           // ******************************************************************************************************
       2: // Start Movement via Processchannel
           // Mode 04 hex = Profile Velocity (RefA32 = target velocity / RefB32 = reserved)
           #ILx2T_Ref.q_dw_refB_32 := 0;
           #ILx2T_Ref.q_dw_refA_16 := INT_TO_WORD(#i_inTargetVelocity);
           #inTargetVelocityHelper := #i_inTargetVelocity;
           #ILx2T_Ref.q_wo_dmControl := #ILx2T_Ref.q_wo_dmControl AND 16#FF80;
           #ILx2T_Ref.q_wo_dmControl := #ILx2T_Ref.q_wo_dmControl OR 16#0004;
           #inState := #inState + 1;
           // ******************************************************************************************************
       3: // Mode Toggle
           #xModeToggleHelper := NOT #ILx2T_Ref.st_ModeStatus.ModeToggle;   // save toggle bit 
           IF NOT #xModeToggleHelper THEN
               #ILx2T_Ref.q_wo_dmControl := #ILx2T_Ref.q_wo_dmControl AND 16#FF7F;
           ELSE
               #ILx2T_Ref.q_wo_dmControl := #ILx2T_Ref.q_wo_dmControl OR 16#0080;
           END_IF;
           #inState := #inState + 1;
           // ******************************************************************************************************
       4: // Check for mode response OK
           // Check for mode toggle and number of operating mode OK
           IF NOT (#xModeToggleHelper XOR #ILx2T_Ref.st_ModeStatus.ModeToggle) AND (#ILx2T_Ref.by_OP_ModeAct = 16#0004) THEN                            // Check operating mode number
               #TON_Timeout(IN := FALSE,
                            PT := t#1s);
               #inState := #inState + 1;
           ELSE
               // TIMEOUT ERROR
               #TON_Timeout(IN := TRUE,
                            PT := t#1s);
               IF #TON_Timeout.Q THEN
                   #TON_Timeout(IN := FALSE,
                                PT := t#1s);
                   #q_xError := TRUE;
                   #inErrorState := #inState;
                   #inState := 100;
               END_IF;
           END_IF;
           // ******************************************************************************************************
       5: // Check operating mode
           // Check for target reached (Drive status x_Add)
           IF (#ILx2T_Ref.i_woDriveStatus AND 16#2000) = 16#2000 THEN  // x_Add = Target vel reached     
               #q_xTargetVelocityReached := TRUE;
           ELSE
               #q_xTargetVelocityReached := FALSE;
           END_IF;
           // x_Error
           IF (#ILx2T_Ref.i_woDriveStatus AND 16#8000) = 16#8000 THEN  // error     
               #inErrorState := #inState;
               #inState := 100;
           // Monitoring of actual operating mode
           ELSIF (#ILx2T_Ref.by_OP_ModeAct <> 16#0004) THEN
               #q_xCommandAborted := TRUE;
               #q_xBusy := FALSE;
               #q_xTargetVelocityReached := FALSE;
               #inState := 110;
           // Check for new target velocity value !
           ELSIF #inTargetVelocityHelper <> #i_inTargetVelocity THEN
               #inState := 2;
           // Check for ABORT command
           ELSIF #i_xAbort THEN
               #ILx2T_Ref.x_QuickStopInt := TRUE;
               #inState := #inState + 1;
           END_IF;
       6:
           #TON_Timeout(IN := TRUE,
                        PT := t#10s);
           IF #TON_Timeout.Q THEN
               #TON_Timeout(IN := FALSE,
                            PT := t#1s);
               #ILx2T_Ref.x_QuickStopInt := FALSE;
               #ILx2T_Ref.x_FaultResetInt := FALSE;
               #q_xError := TRUE;
               #inErrorState := #inState;
               #inState := 100;
           ELSIF #ILx2T_Ref.stDriveStatus.x_End AND (#ILx2T_Ref.i_woDriveStatus AND 16#F) >= 7 THEN  // Check for STANDSTILL
               #ILx2T_Ref.x_QuickStopInt := FALSE;
               #ILx2T_Ref.x_FaultResetInt := TRUE;
           ELSIF #ILx2T_Ref.stDriveStatus.x_End AND (#ILx2T_Ref.i_woDriveStatus AND 16#F) < 7 THEN  // Check for STANDSTILL
               #TON_Timeout(IN := FALSE,
                            PT := t#1s);
               #ILx2T_Ref.x_QuickStopInt := FALSE;
               #ILx2T_Ref.x_FaultResetInt := FALSE;
               #q_xCommandAborted := TRUE;
               #q_xBusy := FALSE;
               #q_xTargetVelocityReached := FALSE;
               #inState := 110;
           END_IF;

           // ******************************************************************************************************
       100:  // Error state
           #q_xBusy := FALSE;
           #q_xError := TRUE;
           #inState := 110;
           // ******************************************************************************************************
       110:  // finished
           IF NOT #i_xExecute AND NOT #i_xAbort THEN
               #q_xTargetVelocityReached := FALSE;
               #q_xError := FALSE;
               #q_xBusy := FALSE;
               #q_xCommandAborted := FALSE;
               #inState := 0;
           END_IF;
           // ******************************************************************************************************
   END_CASE;
END_FUNCTION_BLOCK

FUNCTION_BLOCK "ILx2_ModbusTCP_Data_1500"   // FB10, SCL
{ S7_Optimized_Access := 'FALSE' }
VERSION : 1.5
   VAR_INPUT
      CONNECT_ID_1 : Conn_Ouc := 1;   // unique connection ID DPL Read
      CONNECT_ID_2 : Conn_Ouc := 2;   // unique connection ID DPL Write
      CONNECT_ID_3 : Conn_Ouc := 3;   // unique connection ID Parameter read
      CONNECT_ID_4 : Conn_Ouc := 4;   // unique connection ID Parameter write
      IP_OCTET_1 : USInt := 192;
      IP_OCTET_2 : USInt := 168;
      IP_OCTET_3 : USInt;
      IP_OCTET_4 : USInt;
      inNodeGuardTime : UInt := 1000;   // Modbus Node Guard Time (Object 6544 Range 0..10000 ms)
   END_VAR
   VAR_OUTPUT
      Com_OK : Bool;   // Communication OK
      Error : Bool;   // Communication error
      ErrorCode : Word;   // MB_CLIENT - error code
   END_VAR
   VAR_IN_OUT
      ILx2T_Ref : "ILx2T_Ref";
   END_VAR
   VAR
      ReadData_DPL : Array[0..7] of Byte;   // Read Data Drive Profile Lexium
      WriteData_DPL : Array[0..7] of Byte;   // Write Data Drive Profile Lexium
      ParaRead_Value : DInt;   // Parameter Read Data
      ParaWrite_Value : DInt;   // Parameter Write Data
      iState_Read_DPL : Int;
      iState_Write_DPL : Int;
      iState_Read_Para : Int;
      iState_Write_Para : Int;
      MB_CLIENT_Instance_DPL_Read : MB_CLIENT;
      MB_CLIENT_Instance_DPL_Write : MB_CLIENT;
      MB_CLIENT_Instance_ParaRead : MB_CLIENT;
      MB_CLIENT_Instance_ParaWrite : MB_CLIENT;
      stCONNECT_DPL_Read : TCON_IP_v4;
      stCONNECT_DPL_Write : TCON_IP_v4;
      stCONNECT_Parameter_Read : TCON_IP_v4;
      stCONNECT_Parameter_Write : TCON_IP_v4;
      Index : Int;
      inIndex : Int;
      xNodeGuardInitOK : Bool;
      xErrorReadDPL : Bool;
      xErrorWriteDPL : Bool;
      xErrorReadParameter : Bool;
      xErrorWriteParameter : Bool;
      diErrorCounter_DPL_Read : DInt;
      diErrorCounter_DPL_Write : DInt;
      diErrorCounter_Para_Read : DInt;
      diErrorCounter_Para_Write : DInt;
      woReadDPL_ErrorID : Word;
      woWriteDPL_ErrorID : Word;
      woReadParameter_ErrorID : Word;
      woWriteParameter_ErrorID : Word;
      iStateTimeReadDPL : Int;
      iStateTimeWriteDPL : Int;
      T_ReadDPL : TON_TIME;
      t_ReadDPL_Min : Time := t#5m;
      t_ReadDPL_Act : Time;
      t_ReadDPL_Max : Time;
      T_WriteDPL : TON_TIME;
      t_WriteDPL_Min : Time := t#5m;
      t_WriteDPL_Act : Time;
      t_WriteDPL_Max : Time;
      MB_CLIENT_Instance : MB_CLIENT;
   END_VAR
BEGIN
   // THIS FB uses ModbusTCP 5.0 - 04.02.2019
   // OpenUserCommunication must be set to Version 5.1 - 04.02.2019
   // 23.07.2018 - Using 4 connections to increase the performance of the data exchange
   // ***************************************************************************************
   // S7-1x00 - MB_Client Version 5.0
   // PLC IP address 10.209.177.xxx
   // Modbus slave IP Address 10.209.177.xxx
   // ***************************************************************************************
   // Read DPL Data OF 4 WORDS from slave
   // ***************************************************************************************
   #stCONNECT_DPL_Read.ActiveEstablished := TRUE;
   #stCONNECT_DPL_Read.ConnectionType := 11;    // TCP
   #stCONNECT_DPL_Read.ID := #CONNECT_ID_1;
   #stCONNECT_DPL_Read.InterfaceId := 64;    // PROFINET Network
   #stCONNECT_DPL_Read.LocalPort := 0;
   #stCONNECT_DPL_Read.RemotePort := 502;   // 502 See TIA ONLINE HELP
   #stCONNECT_DPL_Read.RemoteAddress.ADDR[1] := #IP_OCTET_1;
   #stCONNECT_DPL_Read.RemoteAddress.ADDR[2] := #IP_OCTET_2;
   #stCONNECT_DPL_Read.RemoteAddress.ADDR[3] := #IP_OCTET_3;
   #stCONNECT_DPL_Read.RemoteAddress.ADDR[4] := #IP_OCTET_4;
   CASE #iState_Read_DPL OF
       0:  // DISCONNECT
           #MB_CLIENT_Instance_DPL_Read(REQ := FALSE,
                                        DISCONNECT := TRUE,
                                        MB_MODE := 0,
                                        MB_DATA_ADDR := 400001 + 6926,
                                        MB_DATA_LEN := 4,
                                        MB_DATA_PTR := #ReadData_DPL,
                                        CONNECT := #stCONNECT_DPL_Read);
           #iState_Read_DPL := #iState_Read_DPL + 1;
       1:  // CONNECT  
           #MB_CLIENT_Instance_DPL_Read(REQ := false,
                                        DISCONNECT := FALSE,
                                        MB_MODE := 0,
                                        MB_DATA_ADDR := 400001 + 6926,
                                        MB_DATA_LEN := 4,
                                        MB_DATA_PTR := #ReadData_DPL,
                                        CONNECT := #stCONNECT_DPL_Read);
           IF #MB_CLIENT_Instance_DPL_Read.Connected AND NOT #MB_CLIENT_Instance_DPL_Read.BUSY THEN
               IF NOT #xNodeGuardInitOK THEN
                   #iState_Read_DPL := 200;
               ELSE
                   #iState_Read_DPL := #iState_Read_DPL + 1;
               END_IF;
           ELSIF #MB_CLIENT_Instance_DPL_Read.ERROR THEN
               #woReadDPL_ErrorID := #MB_CLIENT_Instance_DPL_Read.STATUS;
               #iState_Read_DPL := #iState_Read_DPL + 100;
           END_IF;
       2:  // Check for DONE AND NOT BUSY
           #MB_CLIENT_Instance_DPL_Read(REQ := TRUE,
                                        DISCONNECT := FALSE,
                                        MB_MODE := 0,
                                        MB_DATA_ADDR := 400001 + 6926,
                                        MB_DATA_LEN := 4,
                                        MB_DATA_PTR := #ReadData_DPL,
                                        CONNECT := #stCONNECT_DPL_Read);
           IF #MB_CLIENT_Instance_DPL_Read.DONE AND NOT #MB_CLIENT_Instance_DPL_Read.BUSY THEN
               #xErrorReadDPL := FALSE;
               #woReadDPL_ErrorID := 0;
               FOR #Index := 0 TO 7 DO
                   #ILx2T_Ref.arInputData[#Index] := #ReadData_DPL[#Index];
               END_FOR;
           ELSIF #MB_CLIENT_Instance_DPL_Read.ERROR THEN
               #woReadDPL_ErrorID := #MB_CLIENT_Instance_DPL_Read.STATUS;
               FOR #Index := 0 TO 7 DO
                   #ILx2T_Ref.arInputData[#Index] := 0;
               END_FOR;
               #iState_Read_DPL := #iState_Read_DPL + 100;
           END_IF;
       100..120:  // Error state
           #xErrorReadDPL := TRUE;
           #diErrorCounter_DPL_Read := #diErrorCounter_DPL_Read + 1;
           #MB_CLIENT_Instance_DPL_Read(REQ := FALSE,
                                        DISCONNECT := TRUE,
                                        MB_MODE := 0,
                                        MB_DATA_ADDR := 400001 + 6926,
                                        MB_DATA_LEN := 4,
                                        MB_DATA_PTR := #ReadData_DPL,
                                        CONNECT := #stCONNECT_DPL_Read);
           #iState_Read_DPL := 0;

           // **********************************************************************************************************
           // ***** Set Modbus Nodeguar time after communication is established once ***********************************
           // **********************************************************************************************************
       200:  // CONNECT  
           #ParaWrite_Value := #inNodeGuardTime;
           #MB_CLIENT_Instance_DPL_Read(REQ := FALSE,
                                        DISCONNECT := FALSE,
                                        MB_MODE := 1,
                                        MB_DATA_ADDR := 400001 + 5644,
                                        MB_DATA_LEN := 2,
                                        MB_DATA_PTR := #ParaWrite_Value,
                                        CONNECT := #stCONNECT_DPL_Read);
           IF #MB_CLIENT_Instance_DPL_Read.Connected AND NOT #MB_CLIENT_Instance_DPL_Read.BUSY THEN
               #woReadDPL_ErrorID := 0;
               #iState_Read_DPL := #iState_Read_DPL + 1;
           ELSIF #MB_CLIENT_Instance_DPL_Read.ERROR THEN
               #woReadDPL_ErrorID := #MB_CLIENT_Instance_DPL_Read.STATUS;
               #iState_Read_DPL := 119;
           END_IF;
       201:  // Write Parameter
           #ParaWrite_Value := #inNodeGuardTime;
           #MB_CLIENT_Instance_DPL_Read(REQ := TRUE,
                                        DISCONNECT := FALSE,
                                        MB_MODE := 1,
                                        MB_DATA_ADDR := 400001 + 5644,
                                        MB_DATA_LEN := 2,
                                        MB_DATA_PTR := #ParaWrite_Value,
                                        CONNECT := #stCONNECT_DPL_Read);
           IF #MB_CLIENT_Instance_DPL_Read.DONE AND NOT #MB_CLIENT_Instance_DPL_Read.BUSY THEN
               #woReadDPL_ErrorID := 0;
               #MB_CLIENT_Instance_DPL_Read(REQ := FALSE,
                                            DISCONNECT := FALSE,
                                            MB_MODE := 1,
                                            MB_DATA_ADDR := 400001 + 5644,
                                            MB_DATA_LEN := 2,
                                            MB_DATA_PTR := #ParaWrite_Value,
                                            CONNECT := #stCONNECT_DPL_Read);
               #xNodeGuardInitOK := TRUE;
               #iState_Read_DPL := 0;
           ELSIF #MB_CLIENT_Instance_DPL_Read.ERROR THEN
               #woReadDPL_ErrorID := #MB_CLIENT_Instance_DPL_Read.STATUS;
               #iState_Read_DPL := 120;
           END_IF;

   END_CASE;
   // ***************************************************************************************
   // Write DPL Data OF 4 WORDS to slave
   // ***************************************************************************************
   #stCONNECT_DPL_Write.ActiveEstablished := TRUE;
   #stCONNECT_DPL_Write.ConnectionType := 11;    // TCP
   #stCONNECT_DPL_Write.ID := #CONNECT_ID_2;
   #stCONNECT_DPL_Write.InterfaceId := 64;    // PROFINET Network
   #stCONNECT_DPL_Write.LocalPort := 0;
   #stCONNECT_DPL_Write.RemotePort := 502;   // 502 See TIA ONLINE HELP
   #stCONNECT_DPL_Write.RemoteAddress.ADDR[1] := #IP_OCTET_1;
   #stCONNECT_DPL_Write.RemoteAddress.ADDR[2] := #IP_OCTET_2;
   #stCONNECT_DPL_Write.RemoteAddress.ADDR[3] := #IP_OCTET_3;
   #stCONNECT_DPL_Write.RemoteAddress.ADDR[4] := #IP_OCTET_4;
   CASE #iState_Write_DPL OF
       0:  // DISCONNECT
           #MB_CLIENT_Instance_DPL_Write(REQ := FALSE,
                                         DISCONNECT := TRUE,
                                         MB_MODE := 1,
                                         MB_DATA_ADDR := 400001 + 6922,
                                         MB_DATA_LEN := 4,
                                         MB_DATA_PTR := #ReadData_DPL,
                                         CONNECT := #stCONNECT_DPL_Write);
           #iState_Write_DPL := #iState_Write_DPL + 1;
       1:  // CONNECT  
           #MB_CLIENT_Instance_DPL_Write(REQ := FALSE,
                                         DISCONNECT := FALSE,
                                         MB_MODE := 1,
                                         MB_DATA_ADDR := 400001 + 6922,
                                         MB_DATA_LEN := 4,
                                         MB_DATA_PTR := #WriteData_DPL,
                                         CONNECT := #stCONNECT_DPL_Write);
           IF #MB_CLIENT_Instance_DPL_Write.Connected AND NOT #MB_CLIENT_Instance_DPL_Write.BUSY THEN
               #woWriteDPL_ErrorID := 0;
               #iState_Write_DPL := #iState_Write_DPL + 1;
           ELSIF #MB_CLIENT_Instance_DPL_Write.ERROR THEN
               #woWriteDPL_ErrorID := #MB_CLIENT_Instance_DPL_Write.STATUS;
               #iState_Write_DPL := #iState_Write_DPL + 100;
           END_IF;
       2:  // Write Data
           FOR #Index := 0 TO 7 DO
               #WriteData_DPL[#Index] := #ILx2T_Ref.arOutputData[#Index];
           END_FOR;
           #MB_CLIENT_Instance_DPL_Write(REQ := TRUE,
                                         DISCONNECT := FALSE,
                                         MB_MODE := 1,
                                         MB_DATA_ADDR := 400001 + 6922,
                                         MB_DATA_LEN := 4,
                                         MB_DATA_PTR := #WriteData_DPL,
                                         CONNECT := #stCONNECT_DPL_Write);
           IF #MB_CLIENT_Instance_DPL_Write.DONE AND NOT #MB_CLIENT_Instance_DPL_Write.BUSY THEN
               #woWriteDPL_ErrorID := 0;
               #xErrorWriteDPL := FALSE;
           ELSIF #MB_CLIENT_Instance_DPL_Write.ERROR THEN
               #woWriteDPL_ErrorID := #MB_CLIENT_Instance_DPL_Write.STATUS;
               #iState_Write_DPL := #iState_Write_DPL + 100;
           END_IF;

       100..120:  // Error state
           #xErrorWriteDPL := TRUE;
           #diErrorCounter_DPL_Write := #diErrorCounter_DPL_Write + 1;
           #MB_CLIENT_Instance_DPL_Write(REQ := FALSE,
                                         DISCONNECT := TRUE,
                                         MB_MODE := 1,
                                         MB_DATA_ADDR := 400001 + 6922,
                                         MB_DATA_LEN := 4,
                                         MB_DATA_PTR := #WriteData_DPL,
                                         CONNECT := #stCONNECT_DPL_Write);
           #iState_Write_DPL := 0;
   END_CASE;
   // ***************************************************************************************
   // ReadParameter
   // ***************************************************************************************
   #stCONNECT_Parameter_Read.ActiveEstablished := TRUE;
   #stCONNECT_Parameter_Read.ConnectionType := 11;    // TCP
   #stCONNECT_Parameter_Read.ID := #CONNECT_ID_3;
   #stCONNECT_Parameter_Read.InterfaceId := 64;    // PROFINET Network
   #stCONNECT_Parameter_Read.LocalPort := 0;
   #stCONNECT_Parameter_Read.RemotePort := 502;   // 502 See TIA ONLINE HELP
   #stCONNECT_Parameter_Read.RemoteAddress.ADDR[1] := #IP_OCTET_1;
   #stCONNECT_Parameter_Read.RemoteAddress.ADDR[2] := #IP_OCTET_2;
   #stCONNECT_Parameter_Read.RemoteAddress.ADDR[3] := #IP_OCTET_3;
   #stCONNECT_Parameter_Read.RemoteAddress.ADDR[4] := #IP_OCTET_4;
   CASE #iState_Read_Para OF
       0:  // DISCONNECT
           #MB_CLIENT_Instance_ParaRead(REQ := FALSE,
                                        DISCONNECT := TRUE,
                                        MB_MODE := 0,
                                        MB_DATA_ADDR := 400001 + #ILx2T_Ref.udi_ModbusAddress_Read,
                                        MB_DATA_LEN := 2,
                                        MB_DATA_PTR := #ParaRead_Value,
                                        CONNECT := #stCONNECT_Parameter_Read);
           #iState_Read_Para := #iState_Read_Para + 1;

           // **********************************************************************************************************
           // ***** Reading parameters *********************************************************************************
           // **********************************************************************************************************
       1:  // CONNECT  
           #MB_CLIENT_Instance_ParaRead(REQ := FALSE,
                                        DISCONNECT := FALSE,
                                        MB_MODE := 0,
                                        MB_DATA_ADDR := 400001 + #ILx2T_Ref.udi_ModbusAddress_Read,
                                        MB_DATA_LEN := 2,
                                        MB_DATA_PTR := #ParaRead_Value,
                                        CONNECT := #stCONNECT_Parameter_Read);
           IF #MB_CLIENT_Instance_ParaRead.Connected AND NOT #MB_CLIENT_Instance_ParaRead.BUSY THEN
               #iState_Read_Para := #iState_Read_Para + 1;
           ELSIF #MB_CLIENT_Instance_ParaRead.ERROR THEN
               #woReadParameter_ErrorID := #MB_CLIENT_Instance_ParaRead.STATUS;
               #iState_Read_Para := #iState_Read_Para + 100;
           END_IF;
       2:  // Read Parameter
           IF #ILx2T_Ref.x_CommandReadParameter THEN
               #iState_Read_Para := #iState_Read_Para + 1;
           ELSE
               // #woReadParameter_ErrorID := 0;
               #xErrorReadParameter := FALSE;
           END_IF;
       3:  // Read Parameter  
           IF NOT #ILx2T_Ref.x_CommandReadParameter THEN
               #MB_CLIENT_Instance_ParaRead(REQ := FALSE,
                                            DISCONNECT := FALSE,
                                            MB_MODE := 0,
                                            MB_DATA_ADDR := 400001 + #ILx2T_Ref.udi_ModbusAddress_Read,
                                            MB_DATA_LEN := 2,
                                            MB_DATA_PTR := #ParaRead_Value,
                                            CONNECT := #stCONNECT_Parameter_Read);
               #woReadParameter_ErrorID := 0;
               #ILx2T_Ref.di_ParameterReadValue := 0;
               #ILx2T_Ref.x_StatusReadParameter_OK := FALSE;
               #iState_Read_Para := #iState_Read_Para - 1;
           ELSIF #ILx2T_Ref.x_CommandReadParameter THEN
               #MB_CLIENT_Instance_ParaRead(REQ := TRUE,
                                            DISCONNECT := FALSE,
                                            MB_MODE := 0,
                                            MB_DATA_ADDR := 400001 + #ILx2T_Ref.udi_ModbusAddress_Read,
                                            MB_DATA_LEN := 2,
                                            MB_DATA_PTR := #ParaRead_Value,
                                            CONNECT := #stCONNECT_Parameter_Read);
               IF #MB_CLIENT_Instance_ParaRead.DONE AND NOT #MB_CLIENT_Instance_ParaRead.BUSY THEN
                   #woReadParameter_ErrorID := 0;
                   #xErrorReadParameter := FALSE;
                   #ILx2T_Ref.di_ParameterReadValue := #ParaRead_Value;
                   #ILx2T_Ref.x_StatusReadParameter_OK := TRUE;
               ELSIF #MB_CLIENT_Instance_ParaRead.ERROR THEN
                   #woReadParameter_ErrorID := #MB_CLIENT_Instance_ParaRead.STATUS;
                   #ILx2T_Ref.x_StatusReadParameter_Error := TRUE;
                   #iState_Read_Para := #iState_Read_Para + 100;
               END_IF;
           END_IF;

       100..120:  // Error state
           #xErrorReadParameter := TRUE;
           #diErrorCounter_Para_Read := #diErrorCounter_Para_Read + 1;
           #MB_CLIENT_Instance_ParaRead(REQ := FALSE,
                                        DISCONNECT := TRUE,
                                        MB_MODE := 0,
                                        MB_DATA_ADDR := 400001 + #ILx2T_Ref.udi_ModbusAddress_Read,
                                        MB_DATA_LEN := 2,
                                        MB_DATA_PTR := #ParaRead_Value,
                                        CONNECT := #stCONNECT_Parameter_Read);
           #iState_Read_Para := 0;
   END_CASE;
   // ***************************************************************************************
   // WriteParameter
   // ***************************************************************************************
   #stCONNECT_Parameter_Write.ActiveEstablished := TRUE;
   #stCONNECT_Parameter_Write.ConnectionType := 11;    // TCP
   #stCONNECT_Parameter_Write.ID := #CONNECT_ID_4;
   #stCONNECT_Parameter_Write.InterfaceId := 64;    // PROFINET Network
   #stCONNECT_Parameter_Write.LocalPort := 0;
   #stCONNECT_Parameter_Write.RemotePort := 502;   // 502 See TIA ONLINE HELP
   #stCONNECT_Parameter_Write.RemoteAddress.ADDR[1] := #IP_OCTET_1;
   #stCONNECT_Parameter_Write.RemoteAddress.ADDR[2] := #IP_OCTET_2;
   #stCONNECT_Parameter_Write.RemoteAddress.ADDR[3] := #IP_OCTET_3;
   #stCONNECT_Parameter_Write.RemoteAddress.ADDR[4] := #IP_OCTET_4;
   CASE #iState_Write_Para OF
       0:  // DISCONNECT
           #MB_CLIENT_Instance_ParaWrite(REQ := FALSE,
                                         DISCONNECT := TRUE,
                                         MB_MODE := 1,
                                         MB_DATA_ADDR := 400001 + #ILx2T_Ref.udi_ModbusAddress_Write,
                                         MB_DATA_LEN := 2,
                                         MB_DATA_PTR := #ParaWrite_Value,
                                         CONNECT := #stCONNECT_Parameter_Write);
           #iState_Write_Para := #iState_Write_Para + 1;
       1:  // Write Data
           IF #ILx2T_Ref.x_CommandWriteParameter AND NOT #ILx2T_Ref.x_Status_WriteParameter_OK AND NOT #ILx2T_Ref.x_Status_WriteParameter_Error THEN
               #iState_Write_Para := 2;
           ELSE
               #xErrorWriteParameter := FALSE;
           END_IF;
           // **********************************************************************************************************
           // ***** Writing parameters *********************************************************************************
           // **********************************************************************************************************
       2:  // CONNECT  
           #ParaWrite_Value := #ILx2T_Ref.di_ParameterWriteValue;
           #MB_CLIENT_Instance_ParaWrite(REQ := FALSE,
                                         DISCONNECT := FALSE,
                                         MB_MODE := 1,
                                         MB_DATA_ADDR := 400001 + #ILx2T_Ref.udi_ModbusAddress_Write,
                                         MB_DATA_LEN := 2,
                                         MB_DATA_PTR := #ParaWrite_Value,
                                         CONNECT := #stCONNECT_Parameter_Write);
           IF #MB_CLIENT_Instance_ParaWrite.Connected AND NOT #MB_CLIENT_Instance_ParaWrite.BUSY THEN
               #woWriteParameter_ErrorID := 0;
               #iState_Write_Para := #iState_Write_Para + 1;
           ELSIF #MB_CLIENT_Instance_ParaWrite.ERROR THEN
               #woWriteParameter_ErrorID := #MB_CLIENT_Instance_ParaWrite.STATUS;
               #iState_Write_Para := #iState_Write_Para + 100;
           END_IF;
       3:  // Write Parameter
           #ParaWrite_Value := #ILx2T_Ref.di_ParameterWriteValue;
           #MB_CLIENT_Instance_ParaWrite(REQ := TRUE,
                                         DISCONNECT := FALSE,
                                         MB_MODE := 1,
                                         MB_DATA_ADDR := 400001 + #ILx2T_Ref.udi_ModbusAddress_Write,
                                         MB_DATA_LEN := 2,
                                         MB_DATA_PTR := #ParaWrite_Value,
                                         CONNECT := #stCONNECT_Parameter_Write);
           IF #MB_CLIENT_Instance_ParaWrite.DONE AND NOT #MB_CLIENT_Instance_ParaWrite.BUSY THEN
               #woWriteParameter_ErrorID := 0;
               #xErrorWriteParameter := FALSE;
               #MB_CLIENT_Instance_ParaWrite(REQ := FALSE,
                                             DISCONNECT := FALSE,
                                             MB_MODE := 1,
                                             MB_DATA_ADDR := 400001 + #ILx2T_Ref.udi_ModbusAddress_Write,
                                             MB_DATA_LEN := 2,
                                             MB_DATA_PTR := #ParaWrite_Value,
                                             CONNECT := #stCONNECT_Parameter_Write);
               #ILx2T_Ref.x_Status_WriteParameter_OK := TRUE;
               #iState_Write_Para := 1;
           ELSIF #MB_CLIENT_Instance_ParaWrite.ERROR THEN
               #ILx2T_Ref.x_Status_WriteParameter_Error := TRUE;
               #woWriteParameter_ErrorID := #MB_CLIENT_Instance_ParaWrite.STATUS;
               #iState_Write_Para := #iState_Write_Para + 100;
           END_IF;

       100..120:  // Error state
           #xErrorWriteParameter := TRUE;
           #diErrorCounter_Para_Write := #diErrorCounter_Para_Write + 1;
           #MB_CLIENT_Instance_ParaWrite(REQ := FALSE,
                                         DISCONNECT := TRUE,
                                         MB_MODE := 1,
                                         MB_DATA_ADDR := 400001 + #ILx2T_Ref.udi_ModbusAddress_Write,
                                         MB_DATA_LEN := 2,
                                         MB_DATA_PTR := #ParaWrite_Value,
                                         CONNECT := #stCONNECT_Parameter_Write);
           #iState_Write_Para := 0;

   END_CASE;

   // ********************************************************************************************
   // Communication OK or Error
   // ********************************************************************************************
   IF NOT #xErrorReadDPL AND NOT #xErrorWriteDPL AND NOT #xErrorReadParameter AND NOT #xErrorWriteParameter THEN
       #Com_OK := TRUE;
       #Error := FALSE;
   ELSE
       #Com_OK := FALSE;
       #Error := TRUE;
   END_IF;
   // ********************************************************************************************
   // Time measurements
   // Only for Diagnostic
   // ********************************************************************************************
   CASE #iStateTimeReadDPL OF
       0:
           IF #MB_CLIENT_Instance_DPL_Read.DONE THEN
               #T_ReadDPL(IN := FALSE,
                          PT := t#2m);
               #T_ReadDPL(IN := TRUE,
                          PT := t#2m);
               #iStateTimeReadDPL := #iStateTimeReadDPL + 1;
           END_IF;
       1:
           #T_ReadDPL(IN := TRUE,
                      PT := t#2m);
           IF #MB_CLIENT_Instance_DPL_Read.DONE THEN
               #t_ReadDPL_Act := #T_ReadDPL.ET;
               IF #t_ReadDPL_Act > #t_ReadDPL_Max THEN
                   #t_ReadDPL_Max := #t_ReadDPL_Act;
               ELSIF #t_ReadDPL_Act < #t_ReadDPL_Min THEN
                   #t_ReadDPL_Min := #t_ReadDPL_Act;
               END_IF;
               #T_ReadDPL(IN := FALSE,
                          PT := t#2m);
               #T_ReadDPL(IN := TRUE,
                          PT := t#2m);
           END_IF;
   END_CASE;


   CASE #iStateTimeWriteDPL OF
       0:
           IF #MB_CLIENT_Instance_DPL_Write.DONE THEN
               #T_WriteDPL(IN := FALSE,
                           PT := t#2m);
               #T_WriteDPL(IN := TRUE,
                           PT := t#2m);
               #iStateTimeWriteDPL := #iStateTimeWriteDPL + 1;
           END_IF;
       1:
           #T_WriteDPL(IN := TRUE,
                       PT := t#2m);
           IF #MB_CLIENT_Instance_DPL_Write.DONE THEN
               #t_WriteDPL_Act := #T_WriteDPL.ET;
               IF #t_WriteDPL_Act > #t_WriteDPL_Max THEN
                   #t_WriteDPL_Max := #t_WriteDPL_Act;
               ELSIF #t_WriteDPL_Act < #t_WriteDPL_Min THEN
                   #t_WriteDPL_Min := #t_WriteDPL_Act;
               END_IF;
               #T_WriteDPL(IN := FALSE,
                           PT := t#2m);
               #T_WriteDPL(IN := TRUE,
                           PT := t#2m);
           END_IF;
   END_CASE;
END_FUNCTION_BLOCK

// folder: Subroutine

FUNCTION_BLOCK "GP_OB_Initialize"   // FB2, SCL
TITLE = OB Service flags
{ S7_Optimized_Access := 'TRUE' }
AUTHOR : Cigliutt
FAMILY : GP
VERSION : 1.1
// This FB will provide the following information: 1# OB duration time 2# Timer clock and OS. IMPORTANT!!! This FB must be initialized each OB100 call, and must be called for each OB!
   VAR_INPUT
      IN_xInitialize : Bool;   // Initialize values (OB100 call)
   END_VAR
   VAR
      STC_rlLastExecValue_s : LReal;   // Last execution tick value [s]
      STC_rlReminder_s : Real;   // Reminder from last execution [ms]
      STC_dElapsed_100ms_ms : DInt;   // Elapsed time for 0.1s
      STC_dElapsed_200ms_ms : DInt;   // Elapsed time for 0.2s
      STC_dElapsed_400ms_ms : DInt;   // Elapsed time for 0.4s
      STC_dElapsed_500ms_ms : DInt;   // Elapsed time for 0.5s
      STC_dElapsed_800ms_ms : DInt;   // Elapsed time for 0.8s
      STC_dElapsed_1s_ms : DInt;   // Elapsed time for 1s
      STC_dElapsed_2s_ms : DInt;   // Elapsed time for 2s
      STC_dElapsed_5s_ms : DInt;   // Elapsed time for 5s
      STC_dElapsed_10s_ms : DInt;   // Elapsed time for 10s
      STC_dElapsed_30s_ms : DInt;   // Elapsed time for 30s
      STC_dElapsed_1min_ms : DInt;   // Elapsed time for 1min
      STC_dElapsed_2min_ms : DInt;   // Elapsed time for 2min
      STC_dElapsed_10min_ms : DInt;   // Elapsed time for 10min
      STC_dElapsed_30min_ms : DInt;   // Elapsed time for 30min
      STC_dElapsed_1h_ms : DInt;   // Elapsed time for 1h
      OUT_dExecutionTime_ms : DInt;   // OB Execution time [ms]
      OUT_dMinExecutionTime_ms : DInt;   // OB Maximum execution time [ms]
      OUT_dMaxExecutionTime_ms : DInt;   // OB Minimum execution time [ms]
      OUT_xOs_100ms : Bool;   // OS each 100ms
      OUT_xOs_200ms : Bool;   // OS each 200ms
      OUT_xOs_400ms : Bool;   // OS each 400ms
      OUT_xOs_500ms : Bool;   // OS each 500ms
      OUT_xOs_800ms : Bool;   // OS each 800ms
      OUT_xOs_1s : Bool;   // OS each 1s
      OUT_xOs_2s : Bool;   // OS each 2s
      OUT_xOs_5s : Bool;   // OS each 5s
      OUT_xOs_10s : Bool;   // OS each 10s
      OUT_xOs_30s : Bool;   // OS each 30s
      OUT_xOs_1min : Bool;   // OS each 1min
      OUT_xOs_2min : Bool;   // OS each 2min
      OUT_xOs_10min : Bool;   // OS each 10min
      OUT_xOs_30min : Bool;   // OS each 30min
      OUT_xOs_1h : Bool;   // OS each 1h
      OUT_xClock_100ms : Bool;   // Clock 100ms
      OUT_xClock_200ms : Bool;   // Clock 200ms
      OUT_xClock_400ms : Bool;   // Clock 400ms
      OUT_xClock_500ms : Bool;   // Clock 500ms
      OUT_xClock_800ms : Bool;   // Clock 800ms
      OUT_xClock_1s : Bool;   // Clock 1s
      OUT_xClock_2s : Bool;   // Clock 2s
      OUT_xClock_5s : Bool;   // Clock 5s
      OUT_xClock_10s : Bool;   // Clock 10s
      OUT_xClock_30s : Bool;   // Clock 30s
      OUT_xClock_1min : Bool;   // Clock 1min
      OUT_xClock_2min : Bool;   // Clock 2min
      OUT_xClock_10min : Bool;   // Clock 10min
      OUT_xClock_30min : Bool;   // Clock 30min
      OUT_xClock_1h : Bool;   // Clock 1h
      OUT_xDebugOFF : Bool;   // Commisioning bit - Always OFF
      OUT_xDebugON : Bool;   // Commisioning bit - Always ON
   END_VAR
   VAR_TEMP
      TMP_rlActualExecutionTime : Real;   // ActualExecutionTime [ms]
      TMP_rlActualExecutionTimeRound : Real;   // Rounded execution time [ms]
      TMP_rlActualExecutionTimeCalculated : Real;
   END_VAR
   VAR CONSTANT
      CONST_DTICK_100MS : DInt := 100;
      CONST_DTICK_200MS : DInt := 200;
      CONST_DTICK_400MS : DInt := 400;
      CONST_DTICK_500MS : DInt := 500;
      CONST_DTICK_800MS : DInt := 800;
      CONST_DTICK_1S : DInt := 1000;
      CONST_DTICK_2S : DInt := 2000;
      CONST_DTICK_5S : DInt := 5000;
      CONST_DTICK_10S : DInt := 10000;
      CONST_DTICK_30S : DInt := 30000;
      CONST_DTICK_1MIN : DInt := 60000;
      CONST_DTICK_2MIN : DInt := 120000;
      CONST_DTICK_10MIN : DInt := 600000;
      CONST_DTICK_30MIN : DInt := 1800000;
      CONST_DTICK_1H : DInt := 86400000;
      CONST_DMAX_INT : DInt := 16#7FFF_FFFF;
   END_VAR
BEGIN
   //Initialize OS bits
   #OUT_xOs_100ms := false;
   #OUT_xOs_200ms := false;
   #OUT_xOs_400ms := false;
   #OUT_xOs_500ms := false;
   #OUT_xOs_800ms := false;
   #OUT_xOs_1s := false;
   #OUT_xOs_2s := false;
   #OUT_xOs_5s := false;
   #OUT_xOs_10s := false;
   #OUT_xOs_30s := false;
   #OUT_xOs_1min := false;
   #OUT_xOs_2min := false;
   #OUT_xOs_10min := false;
   #OUT_xOs_30min := false;
   #OUT_xOs_1h := false;

   //Initialize FB execution
   IF #IN_xInitialize = true THEN


       #IN_xInitialize := false;

       #OUT_dExecutionTime_ms := 0;
       #OUT_dMinExecutionTime_ms := #CONST_DMAX_INT;
       #OUT_dMaxExecutionTime_ms := 0;
       #OUT_xClock_100ms := false;
       #OUT_xClock_200ms := false;
       #OUT_xClock_400ms := false;
       #OUT_xClock_500ms := false;
       #OUT_xClock_800ms := false;
       #OUT_xClock_1s := false;
       #OUT_xClock_2s := false;
       #OUT_xClock_5s := false;
       #OUT_xClock_10s := false;
       #OUT_xClock_30s := false;
       #OUT_xClock_1min := false;
       #OUT_xClock_2min := false;
       #OUT_xClock_10min := false;
       #OUT_xClock_30min := false;
       #OUT_xClock_1h := false;

       #STC_dElapsed_100ms_ms := 0;
       #STC_dElapsed_200ms_ms := 0;
       #STC_dElapsed_400ms_ms := 0;
       #STC_dElapsed_500ms_ms := 0;
       #STC_dElapsed_800ms_ms := 0;
       #STC_dElapsed_1s_ms := 0;
       #STC_dElapsed_2s_ms := 0;
       #STC_dElapsed_5s_ms := 0;
       #STC_dElapsed_10s_ms := 0;
       #STC_dElapsed_30s_ms := 0;
       #STC_dElapsed_1min_ms := 0;
       #STC_dElapsed_2min_ms := 0;
       #STC_dElapsed_10min_ms := 0;
       #STC_dElapsed_30min_ms := 0;
       #STC_dElapsed_1h_ms := 0;
       #STC_rlLastExecValue_s := 0;

   END_IF;
   //***** CALCULATE OB EXECUTION TIME ***** 
   //Take the execution time from the CPU
   #TMP_rlActualExecutionTime := LREAL_TO_REAL(RUNTIME(MEM := #STC_rlLastExecValue_s));

   //Convert from [s] to [ms]
   #TMP_rlActualExecutionTime := #TMP_rlActualExecutionTime * 1000.0;

   //Add the reminder of the last cycle
   #TMP_rlActualExecutionTimeCalculated := #TMP_rlActualExecutionTime + #STC_rlReminder_s;
   //Calculate the rounded value
   #TMP_rlActualExecutionTimeRound := ROUND_REAL(#TMP_rlActualExecutionTimeCalculated);
   #OUT_dExecutionTime_ms := ROUND_DINT(#TMP_rlActualExecutionTimeCalculated);

   //Save the reminder for the next cycle
   #STC_rlReminder_s := #TMP_rlActualExecutionTimeCalculated - #TMP_rlActualExecutionTimeRound;

   //Save the maximum scan value
   IF #OUT_dExecutionTime_ms > #OUT_dMaxExecutionTime_ms THEN
       #OUT_dMaxExecutionTime_ms := #OUT_dExecutionTime_ms;
   END_IF;

   //Save the minimum scan value
   IF #OUT_dExecutionTime_ms < #OUT_dMinExecutionTime_ms THEN
       #OUT_dMinExecutionTime_ms := #OUT_dExecutionTime_ms;
   END_IF;

   //***** CALCULATE SERVICES CLOCK *****

   //Increment counters for each clock
   #STC_dElapsed_100ms_ms := #STC_dElapsed_100ms_ms + #OUT_dExecutionTime_ms;
   #STC_dElapsed_200ms_ms := #STC_dElapsed_200ms_ms + #OUT_dExecutionTime_ms;
   #STC_dElapsed_400ms_ms := #STC_dElapsed_400ms_ms + #OUT_dExecutionTime_ms;
   #STC_dElapsed_500ms_ms := #STC_dElapsed_500ms_ms + #OUT_dExecutionTime_ms;
   #STC_dElapsed_800ms_ms := #STC_dElapsed_800ms_ms + #OUT_dExecutionTime_ms;
   #STC_dElapsed_1s_ms := #STC_dElapsed_1s_ms + #OUT_dExecutionTime_ms;
   #STC_dElapsed_2s_ms := #STC_dElapsed_2s_ms + #OUT_dExecutionTime_ms;
   #STC_dElapsed_5s_ms := #STC_dElapsed_5s_ms + #OUT_dExecutionTime_ms;
   #STC_dElapsed_10s_ms := #STC_dElapsed_10s_ms + #OUT_dExecutionTime_ms;
   #STC_dElapsed_30s_ms := #STC_dElapsed_30s_ms + #OUT_dExecutionTime_ms;
   #STC_dElapsed_1min_ms := #STC_dElapsed_1min_ms + #OUT_dExecutionTime_ms;
   #STC_dElapsed_2min_ms := #STC_dElapsed_2min_ms + #OUT_dExecutionTime_ms;
   #STC_dElapsed_10min_ms := #STC_dElapsed_10min_ms + #OUT_dExecutionTime_ms;
   #STC_dElapsed_30min_ms := #STC_dElapsed_30min_ms + #OUT_dExecutionTime_ms;
   #STC_dElapsed_1h_ms := #STC_dElapsed_1h_ms + #OUT_dExecutionTime_ms;

   //Calculate the 100ms
   IF #STC_dElapsed_100ms_ms >= #CONST_DTICK_100MS THEN
       #STC_dElapsed_100ms_ms := #STC_dElapsed_100ms_ms - #CONST_DTICK_100MS;

       #OUT_xOs_100ms := true;

       IF (#OUT_xClock_100ms = false) THEN
           #OUT_xClock_100ms := true;
       ELSE
           #OUT_xClock_100ms := false;
       END_IF;
   END_IF;

   //Calculate the 200ms
   IF #STC_dElapsed_200ms_ms >= #CONST_DTICK_200MS THEN
       #STC_dElapsed_200ms_ms := #STC_dElapsed_200ms_ms - #CONST_DTICK_200MS;

       #OUT_xOs_200ms := true;

       IF (#OUT_xClock_200ms = false) THEN
           #OUT_xClock_200ms := true;
       ELSE
           #OUT_xClock_200ms := false;
       END_IF;
   END_IF;

   //Calculate the 400ms
   IF #STC_dElapsed_400ms_ms >= #CONST_DTICK_400MS THEN
       #STC_dElapsed_400ms_ms := #STC_dElapsed_400ms_ms - #CONST_DTICK_400MS;

       #OUT_xOs_400ms := true;

       IF (#OUT_xClock_400ms = false) THEN
           #OUT_xClock_400ms := true;
       ELSE
           #OUT_xClock_400ms := false;
       END_IF;
   END_IF;

   //Calculate the 500ms
   IF #STC_dElapsed_500ms_ms >= #CONST_DTICK_500MS THEN
       #STC_dElapsed_500ms_ms := #STC_dElapsed_500ms_ms - #CONST_DTICK_500MS;

       #OUT_xOs_500ms := true;

       IF (#OUT_xClock_500ms = false) THEN
           #OUT_xClock_500ms := true;
       ELSE
           #OUT_xClock_500ms := false;
       END_IF;
   END_IF;

   //Calculate the 800ms
   IF #STC_dElapsed_800ms_ms >= #CONST_DTICK_800MS THEN
       #STC_dElapsed_800ms_ms := #STC_dElapsed_800ms_ms - #CONST_DTICK_800MS;

       #OUT_xOs_800ms := true;

       IF (#OUT_xClock_800ms = false) THEN
           #OUT_xClock_800ms := true;
       ELSE
           #OUT_xClock_800ms := false;
       END_IF;
   END_IF;

   //Calculate the 1s
   IF #STC_dElapsed_1s_ms >= #CONST_DTICK_1S THEN
       #STC_dElapsed_1s_ms := #STC_dElapsed_1s_ms - #CONST_DTICK_1S;

       #OUT_xOs_1s := true;

       IF (#OUT_xClock_1s = false) THEN
           #OUT_xClock_1s := true;
       ELSE
           #OUT_xClock_1s := false;
       END_IF;
   END_IF;

   //Calculate the 2s
   IF #STC_dElapsed_2s_ms >= #CONST_DTICK_2S THEN
       #STC_dElapsed_2s_ms := #STC_dElapsed_2s_ms - #CONST_DTICK_2S;

       #OUT_xOs_2s := true;

       IF (#OUT_xClock_2s = false) THEN
           #OUT_xClock_2s := true;
       ELSE
           #OUT_xClock_2s := false;
       END_IF;
   END_IF;

   //Calculate the 5s
   IF #STC_dElapsed_5s_ms >= #CONST_DTICK_5S THEN
       #STC_dElapsed_5s_ms := #STC_dElapsed_5s_ms - #CONST_DTICK_5S;

       #OUT_xOs_5s := true;

       IF (#OUT_xClock_5s = false) THEN
           #OUT_xClock_5s := true;
       ELSE
           #OUT_xClock_5s := false;
       END_IF;
   END_IF;

   //Calculate the 10s
   IF #STC_dElapsed_10s_ms >= #CONST_DTICK_10S THEN
       #STC_dElapsed_10s_ms := #STC_dElapsed_10s_ms - #CONST_DTICK_10S;

       #OUT_xOs_10s := true;

       IF (#OUT_xClock_10s = false) THEN
           #OUT_xClock_10s := true;
       ELSE
           #OUT_xClock_10s := false;
       END_IF;
   END_IF;

   //Calculate the 30s
   IF #STC_dElapsed_30s_ms >= #CONST_DTICK_30S THEN
       #STC_dElapsed_30s_ms := #STC_dElapsed_30s_ms - #CONST_DTICK_30S;

       #OUT_xOs_30s := true;

       IF (#OUT_xClock_30s = false) THEN
           #OUT_xClock_30s := true;
       ELSE
           #OUT_xClock_30s := false;
       END_IF;
   END_IF;

   //Calculate the 1min
   IF #STC_dElapsed_1min_ms >= #CONST_DTICK_1MIN THEN
       #STC_dElapsed_1min_ms := #STC_dElapsed_1min_ms - #CONST_DTICK_1MIN;

       #OUT_xOs_1min := true;

       IF (#OUT_xClock_1min = false) THEN
           #OUT_xClock_1min := true;
       ELSE
           #OUT_xClock_1min := false;
       END_IF;
   END_IF;

   //Calculate the 2min
   IF #STC_dElapsed_2min_ms >= #CONST_DTICK_2MIN THEN
       #STC_dElapsed_2min_ms := #STC_dElapsed_2min_ms - #CONST_DTICK_2MIN;

       #OUT_xOs_2min := true;

       IF (#OUT_xClock_2min = false) THEN
           #OUT_xClock_2min := true;
       ELSE
           #OUT_xClock_2min := false;
       END_IF;
   END_IF;

   //Calculate the 10min
   IF #STC_dElapsed_10min_ms >= #CONST_DTICK_10MIN THEN
       #STC_dElapsed_10min_ms := #STC_dElapsed_10min_ms - #CONST_DTICK_10MIN;

       #OUT_xOs_10min := true;

       IF (#OUT_xClock_10min = false) THEN
           #OUT_xClock_10min := true;
       ELSE
           #OUT_xClock_10min := false;
       END_IF;
   END_IF;

   //Calculate the 30min
   IF #STC_dElapsed_30min_ms >= #CONST_DTICK_30MIN THEN
       #STC_dElapsed_30min_ms := #STC_dElapsed_30min_ms - #CONST_DTICK_30MIN;

       #OUT_xOs_30min := true;

       IF (#OUT_xClock_30min = false) THEN
           #OUT_xClock_30min := true;
       ELSE
           #OUT_xClock_30min := false;
       END_IF;
   END_IF;

   //Calculate the 1h
   IF #STC_dElapsed_1h_ms >= #CONST_DTICK_1H THEN
       #STC_dElapsed_1h_ms := #STC_dElapsed_1h_ms - #CONST_DTICK_1H;

       #OUT_xOs_1h := true;

       IF (#OUT_xClock_1h = false) THEN
           #OUT_xClock_1h := true;
       ELSE
           #OUT_xClock_1h := false;
       END_IF;
   END_IF;
END_FUNCTION_BLOCK

FUNCTION "GP_GetArraySize" : Int   // FC9, SCL
{ S7_Optimized_Access := 'TRUE' }
AUTHOR : Cigliutt
FAMILY : GP
VERSION : 1.0
   VAR_IN_OUT
      INO_vArray : Variant;
   END_VAR
   VAR_TEMP
      TMP_udNumEl : UDInt;
   END_VAR
BEGIN
   #TMP_udNumEl := 0;

   IF IS_ARRAY(#INO_vArray) THEN
       #TMP_udNumEl := CountOfElements(#INO_vArray);
   END_IF;

   #GP_GetArraySize := UDINT_TO_INT(#TMP_udNumEl);
END_FUNCTION

FUNCTION "GP_BlockMoveStruct" : Int   // FC13, SCL
{ S7_Optimized_Access := 'TRUE' }
AUTHOR : Cigliutt
FAMILY : GP